   1118: 'GCU_ALARM_WORD_08_BIT_14', class GCU Alarms, trigger "60_Alarm_Data_GCU_ALARM_WORD_08" bit 6
   1119: 'GCU_ALARM_WORD_08_BIT_15', class GCU Alarms, trigger "60_Alarm_Data_GCU_ALARM_WORD_08" bit 7
   1120: 'GCU_ALARM_WORD_08_BIT_0', class GCU Alarms, trigger "60_Alarm_Data_GCU_ALARM_WORD_08" bit 8
   1121: 'GCU_ALARM_WORD_08_BIT_1', class GCU Alarms, trigger "60_Alarm_Data_GCU_ALARM_WORD_08" bit 9
   1122: 'GCU_ALARM_WORD_08_BIT_2', class GCU Alarms, trigger "60_Alarm_Data_GCU_ALARM_WORD_08" bit 10
   1123: 'GCU_ALARM_WORD_08_BIT_3', class GCU Alarms, trigger "60_Alarm_Data_GCU_ALARM_WORD_08" bit 11
   1124: 'GCU_ALARM_WORD_08_BIT_4', class GCU Alarms, trigger "60_Alarm_Data_GCU_ALARM_WORD_08" bit 12
   1125: 'GCU_ALARM_WORD_08_BIT_5', class GCU Alarms, trigger "60_Alarm_Data_GCU_ALARM_WORD_08" bit 13
   1126: 'GCU_ALARM_WORD_08_BIT_6', class GCU Alarms, trigger "60_Alarm_Data_GCU_ALARM_WORD_08" bit 14
   1127: 'GCU_ALARM_WORD_08_BIT_7', class GCU Alarms, trigger "60_Alarm_Data_GCU_ALARM_WORD_08" bit 15
   1128: 'GCU_ALARM_WORD_09_BIT_8', class GCU Alarms, trigger "60_Alarm_Data_GCU_ALARM_WORD_09" bit 0
   1129: 'GCU_ALARM_WORD_09_BIT_9', class GCU Alarms, trigger "60_Alarm_Data_GCU_ALARM_WORD_09" bit 1
   1130: 'GCU_ALARM_WORD_09_BIT_10', class GCU Alarms, trigger "60_Alarm_Data_GCU_ALARM_WORD_09" bit 2
   1131: 'GCU_ALARM_WORD_09_BIT_11', class GCU Alarms, trigger "60_Alarm_Data_GCU_ALARM_WORD_09" bit 3
   1132: 'GCU_ALARM_WORD_09_BIT_12', class GCU Alarms, trigger "60_Alarm_Data_GCU_ALARM_WORD_09" bit 4
   1133: 'GCU_ALARM_WORD_09_BIT_13', class GCU Alarms, trigger "60_Alarm_Data_GCU_ALARM_WORD_09" bit 5
   1134: 'GCU_ALARM_WORD_09_BIT_14', class GCU Alarms, trigger "60_Alarm_Data_GCU_ALARM_WORD_09" bit 6
   1135: 'GCU_ALARM_WORD_09_BIT_15', class GCU Alarms, trigger "60_Alarm_Data_GCU_ALARM_WORD_09" bit 7
   1136: 'GCU_ALARM_WORD_09_BIT_0', class GCU Alarms, trigger "60_Alarm_Data_GCU_ALARM_WORD_09" bit 8
   1137: 'GCU_ALARM_WORD_09_BIT_1', class GCU Alarms, trigger "60_Alarm_Data_GCU_ALARM_WORD_09" bit 9
   1138: 'GCU_ALARM_WORD_09_BIT_2', class GCU Alarms, trigger "60_Alarm_Data_GCU_ALARM_WORD_09" bit 10
   1139: 'GCU_ALARM_WORD_09_BIT_3', class GCU Alarms, trigger "60_Alarm_Data_GCU_ALARM_WORD_09" bit 11
   1140: 'GCU_ALARM_WORD_09_BIT_4', class GCU Alarms, trigger "60_Alarm_Data_GCU_ALARM_WORD_09" bit 12
   1141: 'GCU_ALARM_WORD_09_BIT_5', class GCU Alarms, trigger "60_Alarm_Data_GCU_ALARM_WORD_09" bit 13
   1142: 'GCU_ALARM_WORD_09_BIT_6', class GCU Alarms, trigger "60_Alarm_Data_GCU_ALARM_WORD_09" bit 14
   1143: 'GCU_ALARM_WORD_09_BIT_7', class GCU Alarms, trigger "60_Alarm_Data_GCU_ALARM_WORD_09" bit 15
   1144: 'PIT-358 FRESH WATER INLET PRESSURE', class GCU Warnings, trigger "62_Warning_Data_GCU_WARNING_WORD_01" bit 0
   1145: 'GCU_WARNING_WORD_01_BIT_9', class GCU Warnings, trigger "62_Warning_Data_GCU_WARNING_WORD_01" bit 1
   1146: 'GCU_WARNING_WORD_01_BIT_10', class GCU Warnings, trigger "62_Warning_Data_GCU_WARNING_WORD_01" bit 2
   1147: 'GCU_WARNING_WORD_01_BIT_11', class GCU Warnings, trigger "62_Warning_Data_GCU_WARNING_WORD_01" bit 3
   1148: 'GCU_WARNING_WORD_01_BIT_12', class GCU Warnings, trigger "62_Warning_Data_GCU_WARNING_WORD_01" bit 4
   1149: 'GCU_WARNING_WORD_01_BIT_13', class GCU Warnings, trigger "62_Warning_Data_GCU_WARNING_WORD_01" bit 5
   1150: 'GCU_WARNING_WORD_01_BIT_14', class GCU Warnings, trigger "62_Warning_Data_GCU_WARNING_WORD_01" bit 6
   1151: 'GCU_WARNING_WORD_01_BIT_15', class GCU Warnings, trigger "62_Warning_Data_GCU_WARNING_WORD_01" bit 7
   1152: 'PIT-348 CSW PRESSURE - OUT OF RANGE', class GCU Warnings, trigger "62_Warning_Data_GCU_WARNING_WORD_01" bit 8
   1153: 'LIT-304 LIQUID LEVEL - OUT OF RANGE', class GCU Warnings, trigger "62_Warning_Data_GCU_WARNING_WORD_01" bit 9
   1154: 'TIT-406 GAS TO DECK (OUTLET) TEMP - OUT OF RANGE', class GCU Warnings, trigger "62_Warning_Data_GCU_WARNING_WORD_01" bit 10
   1155: 'TIT-408 FRESH WATER COOLING TEMP - OUT OF RANGE', class GCU Warnings, trigger "62_Warning_Data_GCU_WARNING_WORD_01" bit 11
   1156: 'TIT-002 PGC DISCHARGE (OUTLET) TEMP - OUT OF RANGE', class GCU Warnings, trigger "62_Warning_Data_GCU_WARNING_WORD_01" bit 12
   1157: 'PIT-002 PGC DISCHARGE (OUTLET) PRESSURE - OUT OF RANGE', class GCU Warnings, trigger "62_Warning_Data_GCU_WARNING_WORD_01" bit 13
   1158: 'PIT-353 RECIRCULATION FRESH WATER PRESSURE - OUT OF RANGE', class GCU Warnings, trigger "62_Warning_Data_GCU_WARNING_WORD_01" bit 14
   1159: 'PIT-416 GAS TO DECK PRESSURE - OUT OF RANGE', class GCU Warnings, trigger "62_Warning_Data_GCU_WARNING_WORD_01" bit 15
   1160: 'PIT-002 - HIGH', class GCU Warnings, trigger "62_Warning_Data_GCU_WARNING_WORD_02" bit 0
   1161: 'PIT-353 FRESH WATER COOLING TO GCU - LOW', class GCU Warnings, trigger "62_Warning_Data_GCU_WARNING_WORD_02" bit 1
   1162: 'PIT-353 FRESH WATER COOLING TO GCU - HIGH', class GCU Warnings, trigger "62_Warning_Data_GCU_WARNING_WORD_02" bit 2
   1163: 'PIT-416 PROCESS GAS TO DECK PRESSURE - LOW', class GCU Warnings, trigger "62_Warning_Data_GCU_WARNING_WORD_02" bit 3
   1164: 'PIT-416 PROCESS GAS TO DECK PRESSURE - HIGH', class GCU Warnings, trigger "62_Warning_Data_GCU_WARNING_WORD_02" bit 4
   1165: 'PIT-358 BOOSTER FRESH WATER FILL PRESSURE - LOW', class GCU Warnings, trigger "62_Warning_Data_GCU_WARNING_WORD_02" bit 5
   1166: 'PIT-358 BOOSTER FRESH WATER FILL PRESSURE - HIGH', class GCU Warnings, trigger "62_Warning_Data_GCU_WARNING_WORD_02" bit 6
   1167: 'FS-350 FRESH WATER COOLING FLOW SWITCH - LOW FLOW5', class GCU Warnings, trigger "62_Warning_Data_GCU_WARNING_WORD_02" bit 7
   1168: 'CHECK PIT-348 COOLING SEAWATER PRESSURE', class GCU Warnings, trigger "62_Warning_Data_GCU_WARNING_WORD_02" bit 8
   1169: 'CHECK PIT-348 LOW COOLING SEAWATER PRESSURE', class GCU Warnings, trigger "62_Warning_Data_GCU_WARNING_WORD_02" bit 9
   1170: 'CHECK PIT-348 HIGH COOLING SEAWATER PRESSURE', class GCU Warnings, trigger "62_Warning_Data_GCU_WARNING_WORD_02" bit 10
   1171: 'CHECK LIT-304 GCU TANK LEVEL - HIGH', class GCU Warnings, trigger "62_Warning_Data_GCU_WARNING_WORD_02" bit 11
   1172: 'LIT-304 GCU LIQUID LEVEL - LOW', class GCU Warnings, trigger "62_Warning_Data_GCU_WARNING_WORD_02" bit 12
   1173: 'TIT-406 PROCESS GAS TO DECK TEMPERATURE - HIGH TEMP', class GCU Warnings, trigger "62_Warning_Data_GCU_WARNING_WORD_02" bit 13
   1174: 'TIT-408 FRESH WATER COOLING TO GCU TEMPERATURE - HIGH TEMP', class GCU Warnings, trigger "62_Warning_Data_GCU_WARNING_WORD_02" bit 14
   1175: 'CHECK TIT-002 PGC DISCHARGE (OUTLET) TEMPERATURE', class GCU Warnings, trigger "62_Warning_Data_GCU_WARNING_WORD_02" bit 15
   1176: 'GCU_WARNING', class GCU Warnings, trigger "62_Warning_Data_GCU_WARNING_WORD_03" bit 0
   1177: 'GCU_WARNING', class GCU Warnings, trigger "62_Warning_Data_GCU_WARNING_WORD_03" bit 1
   1178: 'GCU_WARNING', class GCU Warnings, trigger "62_Warning_Data_GCU_WARNING_WORD_03" bit 2
   1179: 'GCU_WARNING', class GCU Warnings, trigger "62_Warning_Data_GCU_WARNING_WORD_03" bit 3
   1180: 'GCU_WARNING', class GCU Warnings, trigger "62_Warning_Data_GCU_WARNING_WORD_03" bit 4
   1181: 'GCU_WARNING', class GCU Warnings, trigger "62_Warning_Data_GCU_WARNING_WORD_03" bit 5
   1182: 'GCU_WARNING', class GCU Warnings, trigger "62_Warning_Data_GCU_WARNING_WORD_03" bit 6
   1183: 'GCU_WARNING', class GCU Warnings, trigger "62_Warning_Data_GCU_WARNING_WORD_03" bit 7
   1184: 'LS-303 GCU LIQUID LEVEL - LOW', class GCU Warnings, trigger "62_Warning_Data_GCU_WARNING_WORD_03" bit 8
   1185: 'GCU_WARNING_WORD_03_BIT_1', class GCU Warnings, trigger "62_Warning_Data_GCU_WARNING_WORD_03" bit 9
   1186: 'GCU E-400 - FAULT', class GCU Warnings, trigger "62_Warning_Data_GCU_WARNING_WORD_03" bit 10
   1187: 'TIT-408 FRESH WATER COOLING TO GCU TEMPERATURE - HIGH HIGH TEMP', class GCU Warnings, trigger "62_Warning_Data_GCU_WARNING_WORD_03" bit 11
   1188: 'TIT-406 PROCESS GAS TO DECK TEMPERATURE - HIGH HIGH TEMP', class GCU Warnings, trigger "62_Warning_Data_GCU_WARNING_WORD_03" bit 12
   1189: 'GCU_WARNING_WORD_03_BIT_5', class GCU Warnings, trigger "62_Warning_Data_GCU_WARNING_WORD_03" bit 13
   1190: 'GCU_WARNING_WORD_03_BIT_6', class GCU Warnings, trigger "62_Warning_Data_GCU_WARNING_WORD_03" bit 14
   1191: 'GCU_WARNING_WORD_03_BIT_7', class GCU Warnings, trigger "62_Warning_Data_GCU_WARNING_WORD_03" bit 15
   1192: 'GCU_WARNING_WORD_04_BIT_8', class GCU Warnings, trigger "62_Warning_Data_GCU_WARNING_WORD_04" bit 0
   1193: 'GCU_WARNING_WORD_04_BIT_9', class GCU Warnings, trigger "62_Warning_Data_GCU_WARNING_WORD_04" bit 1
   1194: 'GCU_WARNING_WORD_04_BIT_10', class GCU Warnings, trigger "62_Warning_Data_GCU_WARNING_WORD_04" bit 2
   1195: 'GCU_WARNING_WORD_04_BIT_11', class GCU Warnings, trigger "62_Warning_Data_GCU_WARNING_WORD_04" bit 3
   1196: 'GCU_WARNING_WORD_04_BIT_12', class GCU Warnings, trigger "62_Warning_Data_GCU_WARNING_WORD_04" bit 4
   1197: 'GCU_WARNING_WORD_04_BIT_13', class GCU Warnings, trigger "62_Warning_Data_GCU_WARNING_WORD_04" bit 5
   1198: 'GCU_WARNING_WORD_04_BIT_14', class GCU Warnings, trigger "62_Warning_Data_GCU_WARNING_WORD_04" bit 6
   1199: 'GCU_WARNING_WORD_04_BIT_15', class GCU Warnings, trigger "62_Warning_Data_GCU_WARNING_WORD_04" bit 7
   1200: 'GCU_WARNING_WORD_04_BIT_0', class GCU Warnings, trigger "62_Warning_Data_GCU_WARNING_WORD_04" bit 8
   1201: 'GCU_WARNING_WORD_04_BIT_1', class GCU Warnings, trigger "62_Warning_Data_GCU_WARNING_WORD_04" bit 9
   1202: 'GCU_WARNING_WORD_04_BIT_2', class GCU Warnings, trigger "62_Warning_Data_GCU_WARNING_WORD_04" bit 10
   1203: 'GCU_WARNING_WORD_04_BIT_3', class GCU Warnings, trigger "62_Warning_Data_GCU_WARNING_WORD_04" bit 11
   1204: 'GCU_WARNING_WORD_04_BIT_4', class GCU Warnings, trigger "62_Warning_Data_GCU_WARNING_WORD_04" bit 12
   1205: 'GCU_WARNING_WORD_04_BIT_5', class GCU Warnings, trigger "62_Warning_Data_GCU_WARNING_WORD_04" bit 13
   1206: 'GCU_WARNING_WORD_04_BIT_6', class GCU Warnings, trigger "62_Warning_Data_GCU_WARNING_WORD_04" bit 14
   1207: 'GCU_WARNING_WORD_04_BIT_7', class GCU Warnings, trigger "62_Warning_Data_GCU_WARNING_WORD_04" bit 15
   1208: 'GCU_WARNING_WORD_05_BIT_8', class GCU Warnings, trigger "62_Warning_Data_GCU_WARNING_WORD_05" bit 0
   1209: 'GCU_WARNING_WORD_05_BIT_9', class GCU Warnings, trigger "62_Warning_Data_GCU_WARNING_WORD_05" bit 1
   1210: 'GCU_WARNING_WORD_05_BIT_10', class GCU Warnings, trigger "62_Warning_Data_GCU_WARNING_WORD_05" bit 2
   1211: 'GCU_WARNING_WORD_05_BIT_11', class GCU Warnings, trigger "62_Warning_Data_GCU_WARNING_WORD_05" bit 3
   1212: 'GCU_WARNING_WORD_05_BIT_12', class GCU Warnings, trigger "62_Warning_Data_GCU_WARNING_WORD_05" bit 4
   1213: 'GCU_WARNING_WORD_05_BIT_13', class GCU Warnings, trigger "62_Warning_Data_GCU_WARNING_WORD_05" bit 5
   1214: 'GCU_WARNING_WORD_05_BIT_14', class GCU Warnings, trigger "62_Warning_Data_GCU_WARNING_WORD_05" bit 6
   1215: 'GCU_WARNING_WORD_05_BIT_15', class GCU Warnings, trigger "62_Warning_Data_GCU_WARNING_WORD_05" bit 7
   1216: 'GCU_WARNING_WORD_05_BIT_0', class GCU Warnings, trigger "62_Warning_Data_GCU_WARNING_WORD_05" bit 8
   1217: 'GCU_WARNING_WORD_05_BIT_1', class GCU Warnings, trigger "62_Warning_Data_GCU_WARNING_WORD_05" bit 9
   1218: 'GCU_WARNING_WORD_05_BIT_2', class GCU Warnings, trigger "62_Warning_Data_GCU_WARNING_WORD_05" bit 10
   1219: 'GCU_WARNING_WORD_05_BIT_3', class GCU Warnings, trigger "62_Warning_Data_GCU_WARNING_WORD_05" bit 11
   1220: 'GCU_WARNING_WORD_05_BIT_4', class GCU Warnings, trigger "62_Warning_Data_GCU_WARNING_WORD_05" bit 12
   1221: 'GCU_WARNING_WORD_05_BIT_5', class GCU Warnings, trigger "62_Warning_Data_GCU_WARNING_WORD_05" bit 13
   1222: 'GCU_WARNING_WORD_05_BIT_6', class GCU Warnings, trigger "62_Warning_Data_GCU_WARNING_WORD_05" bit 14
   1223: 'GCU_WARNING_WORD_05_BIT_7', class GCU Warnings, trigger "62_Warning_Data_GCU_WARNING_WORD_05" bit 15
   1224: 'GCU_WARNING_WORD_06_BIT_8', class GCU Warnings, trigger "62_Warning_Data_GCU_WARNING_WORD_06" bit 0
   1225: 'GCU_WARNING_WORD_06_BIT_9', class GCU Warnings, trigger "62_Warning_Data_GCU_WARNING_WORD_06" bit 1
   1226: 'GCU_WARNING_WORD_06_BIT_10', class GCU Warnings, trigger "62_Warning_Data_GCU_WARNING_WORD_06" bit 2
   1227: 'GCU_WARNING_WORD_06_BIT_11', class GCU Warnings, trigger "62_Warning_Data_GCU_WARNING_WORD_06" bit 3
   1228: 'GCU_WARNING_WORD_06_BIT_12', class GCU Warnings, trigger "62_Warning_Data_GCU_WARNING_WORD_06" bit 4
   1229: 'GCU_WARNING_WORD_06_BIT_13', class GCU Warnings, trigger "62_Warning_Data_GCU_WARNING_WORD_06" bit 5
   1230: 'GCU_WARNING_WORD_06_BIT_14', class GCU Warnings, trigger "62_Warning_Data_GCU_WARNING_WORD_06" bit 6
   1231: 'GCU_WARNING_WORD_06_BIT_15', class GCU Warnings, trigger "62_Warning_Data_GCU_WARNING_WORD_06" bit 7
   1232: 'GCU_WARNING_WORD_06_BIT_0', class GCU Warnings, trigger "62_Warning_Data_GCU_WARNING_WORD_06" bit 8
   1233: 'GCU_WARNING_WORD_06_BIT_1', class GCU Warnings, trigger "62_Warning_Data_GCU_WARNING_WORD_06" bit 9
   1234: 'GCU_WARNING_WORD_06_BIT_2', class GCU Warnings, trigger "62_Warning_Data_GCU_WARNING_WORD_06" bit 10
   1235: 'GCU_WARNING_WORD_06_BIT_3', class GCU Warnings, trigger "62_Warning_Data_GCU_WARNING_WORD_06" bit 11
   1236: 'GCU_WARNING_WORD_06_BIT_4', class GCU Warnings, trigger "62_Warning_Data_GCU_WARNING_WORD_06" bit 12
   1237: 'GCU_WARNING_WORD_06_BIT_5', class GCU Warnings, trigger "62_Warning_Data_GCU_WARNING_WORD_06" bit 13
   1238: 'GCU_WARNING_WORD_06_BIT_6', class GCU Warnings, trigger "62_Warning_Data_GCU_WARNING_WORD_06" bit 14
   1239: 'GCU_WARNING_WORD_06_BIT_7', class GCU Warnings, trigger "62_Warning_Data_GCU_WARNING_WORD_06" bit 15
   1240: 'GCU_WARNING_WORD_07_BIT_8', class GCU Warnings, trigger "62_Warning_Data_GCU_WARNING_WORD_07" bit 0
   1241: 'GCU_WARNING_WORD_07_BIT_9', class GCU Warnings, trigger "62_Warning_Data_GCU_WARNING_WORD_07" bit 1
   1242: 'GCU_WARNING_WORD_07_BIT_10', class GCU Warnings, trigger "62_Warning_Data_GCU_WARNING_WORD_07" bit 2
   1243: 'GCU_WARNING_WORD_07_BIT_11', class GCU Warnings, trigger "62_Warning_Data_GCU_WARNING_WORD_07" bit 3
   1244: 'GCU_WARNING_WORD_07_BIT_12', class GCU Warnings, trigger "62_Warning_Data_GCU_WARNING_WORD_07" bit 4
   1245: 'GCU_WARNING_WORD_07_BIT_13', class GCU Warnings, trigger "62_Warning_Data_GCU_WARNING_WORD_07" bit 5
   1246: 'GCU_WARNING_WORD_07_BIT_14', class GCU Warnings, trigger "62_Warning_Data_GCU_WARNING_WORD_07" bit 6
   1247: 'GCU_WARNING_WORD_07_BIT_15', class GCU Warnings, trigger "62_Warning_Data_GCU_WARNING_WORD_07" bit 7
   1248: 'GCU_WARNING_WORD_07_BIT_0', class GCU Warnings, trigger "62_Warning_Data_GCU_WARNING_WORD_07" bit 8
   1249: 'GCU_WARNING_WORD_07_BIT_1', class GCU Warnings, trigger "62_Warning_Data_GCU_WARNING_WORD_07" bit 9
   1250: 'GCU_WARNING_WORD_07_BIT_2', class GCU Warnings, trigger "62_Warning_Data_GCU_WARNING_WORD_07" bit 10
   1251: 'GCU_WARNING_WORD_07_BIT_3', class GCU Warnings, trigger "62_Warning_Data_GCU_WARNING_WORD_07" bit 11
   1252: 'GCU_WARNING_WORD_07_BIT_4', class GCU Warnings, trigger "62_Warning_Data_GCU_WARNING_WORD_07" bit 12
   1253: 'GCU_WARNING_WORD_07_BIT_5', class GCU Warnings, trigger "62_Warning_Data_GCU_WARNING_WORD_07" bit 13
   1254: 'GCU_WARNING_WORD_07_BIT_6', class GCU Warnings, trigger "62_Warning_Data_GCU_WARNING_WORD_07" bit 14
   1255: 'GCU_WARNING_WORD_07_BIT_7', class GCU Warnings, trigger "62_Warning_Data_GCU_WARNING_WORD_07" bit 15
   1256: 'GCU_WARNING_WORD_08_BIT_8', class GCU Warnings, trigger "62_Warning_Data_GCU_WARNING_WORD_08" bit 0
   1257: 'GCU_WARNING_WORD_08_BIT_9', class GCU Warnings, trigger "62_Warning_Data_GCU_WARNING_WORD_08" bit 1
   1258: 'GCU_WARNING_WORD_08_BIT_10', class GCU Warnings, trigger "62_Warning_Data_GCU_WARNING_WORD_08" bit 2
   1259: 'GCU_WARNING_WORD_08_BIT_11', class GCU Warnings, trigger "62_Warning_Data_GCU_WARNING_WORD_08" bit 3
   1260: 'GCU_WARNING_WORD_08_BIT_12', class GCU Warnings, trigger "62_Warning_Data_GCU_WARNING_WORD_08" bit 4
   1261: 'GCU_WARNING_WORD_08_BIT_13', class GCU Warnings, trigger "62_Warning_Data_GCU_WARNING_WORD_08" bit 5
   1262: 'GCU_WARNING_WORD_08_BIT_14', class GCU Warnings, trigger "62_Warning_Data_GCU_WARNING_WORD_08" bit 6
   1263: 'GCU_WARNING_WORD_08_BIT_15', class GCU Warnings, trigger "62_Warning_Data_GCU_WARNING_WORD_08" bit 7
   1264: 'GCU_WARNING_WORD_08_BIT_0', class GCU Warnings, trigger "62_Warning_Data_GCU_WARNING_WORD_08" bit 8
   1265: 'GCU_WARNING_WORD_08_BIT_1', class GCU Warnings, trigger "62_Warning_Data_GCU_WARNING_WORD_08" bit 9
   1266: 'GCU_WARNING_WORD_08_BIT_2', class GCU Warnings, trigger "62_Warning_Data_GCU_WARNING_WORD_08" bit 10
   1267: 'GCU_WARNING_WORD_08_BIT_3', class GCU Warnings, trigger "62_Warning_Data_GCU_WARNING_WORD_08" bit 11
   1268: 'GCU_WARNING_WORD_08_BIT_4', class GCU Warnings, trigger "62_Warning_Data_GCU_WARNING_WORD_08" bit 12
   1269: 'GCU_WARNING_WORD_08_BIT_5', class GCU Warnings, trigger "62_Warning_Data_GCU_WARNING_WORD_08" bit 13
   1270: 'GCU_WARNING_WORD_08_BIT_6', class GCU Warnings, trigger "62_Warning_Data_GCU_WARNING_WORD_08" bit 14
   1271: 'GCU_WARNING_WORD_08_BIT_7', class GCU Warnings, trigger "62_Warning_Data_GCU_WARNING_WORD_08" bit 15
   1272: 'GCU_WARNING_WORD_09_BIT_8', class GCU Warnings, trigger "62_Warning_Data_GCU_WARNING_WORD_09" bit 0
   1273: 'GCU_WARNING_WORD_09_BIT_9', class GCU Warnings, trigger "62_Warning_Data_GCU_WARNING_WORD_09" bit 1
   1274: 'GCU_WARNING_WORD_09_BIT_10', class GCU Warnings, trigger "62_Warning_Data_GCU_WARNING_WORD_09" bit 2
   1275: 'GCU_WARNING_WORD_09_BIT_11', class GCU Warnings, trigger "62_Warning_Data_GCU_WARNING_WORD_09" bit 3
   1276: 'GCU_WARNING_WORD_09_BIT_12', class GCU Warnings, trigger "62_Warning_Data_GCU_WARNING_WORD_09" bit 4
   1277: 'GCU_WARNING_WORD_09_BIT_13', class GCU Warnings, trigger "62_Warning_Data_GCU_WARNING_WORD_09" bit 5
   1278: 'GCU_WARNING_WORD_09_BIT_14', class GCU Warnings, trigger "62_Warning_Data_GCU_WARNING_WORD_09" bit 6
   1279: 'GCU_WARNING_WORD_09_BIT_15', class GCU Warnings, trigger "62_Warning_Data_GCU_WARNING_WORD_09" bit 7
   1280: 'GCU_WARNING_WORD_09_BIT_0', class GCU Warnings, trigger "62_Warning_Data_GCU_WARNING_WORD_09" bit 8
   1281: 'GCU_WARNING_WORD_09_BIT_1', class GCU Warnings, trigger "62_Warning_Data_GCU_WARNING_WORD_09" bit 9
   1282: 'GCU_WARNING_WORD_09_BIT_2', class GCU Warnings, trigger "62_Warning_Data_GCU_WARNING_WORD_09" bit 10
   1283: 'GCU_WARNING_WORD_09_BIT_3', class GCU Warnings, trigger "62_Warning_Data_GCU_WARNING_WORD_09" bit 11
   1284: 'GCU_WARNING_WORD_09_BIT_4', class GCU Warnings, trigger "62_Warning_Data_GCU_WARNING_WORD_09" bit 12
   1285: 'GCU_WARNING_WORD_09_BIT_5', class GCU Warnings, trigger "62_Warning_Data_GCU_WARNING_WORD_09" bit 13
   1286: 'GCU_WARNING_WORD_09_BIT_6', class GCU Warnings, trigger "62_Warning_Data_GCU_WARNING_WORD_09" bit 14
   1287: 'GCU_WARNING_WORD_09_BIT_7', class GCU Warnings, trigger "62_Warning_Data_GCU_WARNING_WORD_09" bit 15
   2000: 'FIT-418 2 PORT USD FLOW - LOW LOW', class Tank Control Alarms, trigger "2060_Alarm_Data_BTCS_ALARM_WORD_01" bit 0
   2001: 'FIT-418 2 PORT USD FLOW - HIGH HIGH', class Tank Control Alarms, trigger "2060_Alarm_Data_BTCS_ALARM_WORD_01" bit 1
   2002: 'FIT-420 2 PORT MBG FLOW - LOW LOW', class Tank Control Alarms, trigger "2060_Alarm_Data_BTCS_ALARM_WORD_01" bit 2
   2003: 'FIT-420 2 PORT MBG FLOW - HIGH HIGH', class Tank Control Alarms, trigger "2060_Alarm_Data_BTCS_ALARM_WORD_01" bit 3
   2004: 'FIT-417 2 STARBOARD USD FLOW - LOW LOW', class Tank Control Alarms, trigger "2060_Alarm_Data_BTCS_ALARM_WORD_01" bit 4
   2005: 'FIT-417 2 STARBOARD USD FLOW - HIGH HIGH', class Tank Control Alarms, trigger "2060_Alarm_Data_BTCS_ALARM_WORD_01" bit 5
   2006: 'FIT-419 2 STARBOARD MBG FLOW - LOW LOW', class Tank Control Alarms, trigger "2060_Alarm_Data_BTCS_ALARM_WORD_01" bit 6
   2007: 'FIT-419 2 STARBOARD MBG FLOW - HIGH HIGH', class Tank Control Alarms, trigger "2060_Alarm_Data_BTCS_ALARM_WORD_01" bit 7
   2008: 'CV-442 2 PORT GAS to TANK VALVE FAULT', class Tank Control Alarms, trigger "2060_Alarm_Data_BTCS_ALARM_WORD_01" bit 8
   2009: 'CV-441 2 STARBOARD GAS to TANK VALVE FAULT', class Tank Control Alarms, trigger "2060_Alarm_Data_BTCS_ALARM_WORD_01" bit 9
   2010: 'TIT-436 2 PORT BWT TEMP - HIGH HIGH', class Tank Control Alarms, trigger "2060_Alarm_Data_BTCS_ALARM_WORD_01" bit 10
   2011: 'TIT-436 2 STARBOARD BWT TEMP - HIGH HIGH', class Tank Control Alarms, trigger "2060_Alarm_Data_BTCS_ALARM_WORD_01" bit 11
   2012: 'LS-425 2 PORT LEVEL - HIGH HIGH', class Tank Control Alarms, trigger "2060_Alarm_Data_BTCS_ALARM_WORD_01" bit 12
   2013: 'LS-425 2 STARBOARD LEVEL - HIGH HIGH', class Tank Control Alarms, trigger "2060_Alarm_Data_BTCS_ALARM_WORD_01" bit 13
   2014: 'PS-436 2 BALLAST TANK PRESSURE - HIGH', class Tank Control Alarms, trigger "2060_Alarm_Data_BTCS_ALARM_WORD_01" bit 14
   2015: '600-TX-433 APT O2 MONITOR - LOW', class Tank Control Alarms, trigger "2060_Alarm_Data_BTCS_ALARM_WORD_01" bit 15
   2016: 'CV422 FPT GAS to TANK VALVE FAULT', class Tank Control Alarms, trigger "2060_Alarm_Data_BTCS_ALARM_WORD_02" bit 0
   2017: 'CV422 1 PORT GAS to TANK VALVE FAULT', class Tank Control Alarms, trigger "2060_Alarm_Data_BTCS_ALARM_WORD_02" bit 1
   2018: 'CV421 1 STARBOARD GAS to TANK VALVE FAULT', class Tank Control Alarms, trigger "2060_Alarm_Data_BTCS_ALARM_WORD_02" bit 2
   2019: 'CV422 3 PORT GAS to TANK VALVE FAULT', class Tank Control Alarms, trigger "2060_Alarm_Data_BTCS_ALARM_WORD_02" bit 3
   2020: 'CV421 3 STARBOARD GAS to TANK VALVE FAULT', class Tank Control Alarms, trigger "2060_Alarm_Data_BTCS_ALARM_WORD_02" bit 4
   2021: 'CV422 4 PORT GAS to TANK VALVE FAULT', class Tank Control Alarms, trigger "2060_Alarm_Data_BTCS_ALARM_WORD_02" bit 5
   2022: 'CV421 4 STARBOARD GAS to TANK VALVE FAULT', class Tank Control Alarms, trigger "2060_Alarm_Data_BTCS_ALARM_WORD_02" bit 6
   2023: 'CV422 5 PORT GAS to TANK VALVE FAULT', class Tank Control Alarms, trigger "2060_Alarm_Data_BTCS_ALARM_WORD_02" bit 7
   2024: 'PIT-415 2 PORT DECK IG PRESSURE - LOW LOW', class Tank Control Alarms, trigger "2060_Alarm_Data_BTCS_ALARM_WORD_02" bit 8
   2025: 'PIT-415 2 PORT DECK IG PRESSURE - HIGH HIGH', class Tank Control Alarms, trigger "2060_Alarm_Data_BTCS_ALARM_WORD_02" bit 9
   2026: 'PIT-415 2 STARBOARD DECK IG PRESSURE - LOW LOW', class Tank Control Alarms, trigger "2060_Alarm_Data_BTCS_ALARM_WORD_02" bit 10
   2027: 'PIT-415 2 STARBOARD DECK IG PRESSURE - HIGH HIGH', class Tank Control Alarms, trigger "2060_Alarm_Data_BTCS_ALARM_WORD_02" bit 11
   2028: 'PIT-424 2 PORT TANK PRESSURE - LOW LOW', class Tank Control Alarms, trigger "2060_Alarm_Data_BTCS_ALARM_WORD_02" bit 12
   2029: 'PIT-424 2 PORT TANK PRESSURE - HIGH HIGH', class Tank Control Alarms, trigger "2060_Alarm_Data_BTCS_ALARM_WORD_02" bit 13
   2030: 'PIT-424 2 STARBOARD TANK PRESSURE - LOW LOW', class Tank Control Alarms, trigger "2060_Alarm_Data_BTCS_ALARM_WORD_02" bit 14
   2031: 'PIT-424 2 STARBOARD TANK PRESSURE - HIGH HIGH', class Tank Control Alarms, trigger "2060_Alarm_Data_BTCS_ALARM_WORD_02" bit 15
   2128: 'FIT-418 2 PORT USD FLOW - LOW', class Tank Control Warnings, trigger "2062_Warning_Data_BTCS_WARNING_WORD_01" bit 0
   2129: 'FIT-418 2 PORT USD FLOW - HIGH', class Tank Control Warnings, trigger "2062_Warning_Data_BTCS_WARNING_WORD_01" bit 1
   2130: 'FIT-420 2 PORT MBG FLOW - LOW', class Tank Control Warnings, trigger "2062_Warning_Data_BTCS_WARNING_WORD_01" bit 2
   2131: 'FIT-420 2 PORT MBG FLOW - HIGH', class Tank Control Warnings, trigger "2062_Warning_Data_BTCS_WARNING_WORD_01" bit 3
   2132: 'FIT-417 2 STARBOARD USD FLOW - LOW', class Tank Control Warnings, trigger "2062_Warning_Data_BTCS_WARNING_WORD_01" bit 4
   2133: 'FIT-417 2 STARBOARD USD FLOW - HIGH', class Tank Control Warnings, trigger "2062_Warning_Data_BTCS_WARNING_WORD_01" bit 5
   2134: 'FIT-419 2 STARBOARD MBG FLOW - LOW', class Tank Control Warnings, trigger "2062_Warning_Data_BTCS_WARNING_WORD_01" bit 6
   2135: 'FIT-419 2 STARBOARD MBG FLOW - HIGH', class Tank Control Warnings, trigger "2062_Warning_Data_BTCS_WARNING_WORD_01" bit 7
   2136: '600-TX-433 APT O2 MONITOR - LOW', class Tank Control Warnings, trigger "2062_Warning_Data_BTCS_WARNING_WORD_01" bit 8
   2137: '600-TX-433 APT O2 MONITOR - LOW LOW', class Tank Control Warnings, trigger "2062_Warning_Data_BTCS_WARNING_WORD_01" bit 9
   2138: 'TIT-436 2 PORT BWT TEMP - HIGH', class Tank Control Warnings, trigger "2062_Warning_Data_BTCS_WARNING_WORD_01" bit 10
   2139: 'TIT-436 2 STARBOARD BWT TEMP - HIGH', class Tank Control Warnings, trigger "2062_Warning_Data_BTCS_WARNING_WORD_01" bit 11
   2140: 'BTCS_WARNING_WORD_01_BIT_4', class Tank Control Warnings, trigger "2062_Warning_Data_BTCS_WARNING_WORD_01" bit 12
   2141: 'BTCS_WARNING_WORD_01_BIT_5', class Tank Control Warnings, trigger "2062_Warning_Data_BTCS_WARNING_WORD_01" bit 13
   2142: 'BTCS_WARNING_WORD_01_BIT_6', class Tank Control Warnings, trigger "2062_Warning_Data_BTCS_WARNING_WORD_01" bit 14
   2143: 'BTCS_WARNING_WORD_01_BIT_7', class Tank Control Warnings, trigger "2062_Warning_Data_BTCS_WARNING_WORD_01" bit 15
   2144: 'TT-426 1 FOR PEACK TANK TEMPERATURE - HIGH', class Tank Control Warnings, trigger "2062_Warning_Data_BTCS_WARNING_WORD_02" bit 0
   2145: 'TT-426 1 PORT TANK TEMPERATURE - HIGH', class Tank Control Warnings, trigger "2062_Warning_Data_BTCS_WARNING_WORD_02" bit 1
   2146: 'TT-426 1 STARBOARD TANK TEMPERATURE - HIGH', class Tank Control Warnings, trigger "2062_Warning_Data_BTCS_WARNING_WORD_02" bit 2
   2147: 'TT-426 3 PORT TANK TEMPERATURE - HIGH', class Tank Control Warnings, trigger "2062_Warning_Data_BTCS_WARNING_WORD_02" bit 3
   2148: 'TT-426 3 STARBOARD TANK TEMPERATURE - HIGH', class Tank Control Warnings, trigger "2062_Warning_Data_BTCS_WARNING_WORD_02" bit 4
   2149: 'TT-426 4 PORT TANK TEMPERATURE - HIGH', class Tank Control Warnings, trigger "2062_Warning_Data_BTCS_WARNING_WORD_02" bit 5
   2150: 'TT-426 4 STARBOARD TANK TEMPERATURE - HIGH', class Tank Control Warnings, trigger "2062_Warning_Data_BTCS_WARNING_WORD_02" bit 6
   2151: 'TT-426 5 PORT TANK TEMPERATURE - HIGH', class Tank Control Warnings, trigger "2062_Warning_Data_BTCS_WARNING_WORD_02" bit 7
   2152: 'PIT-415 2 PORT DECK IG PRESSURE - LOW', class Tank Control Warnings, trigger "2062_Warning_Data_BTCS_WARNING_WORD_02" bit 8
   2153: 'PIT-415 2 PORT DECK IG PRESSURE - HIGH', class Tank Control Warnings, trigger "2062_Warning_Data_BTCS_WARNING_WORD_02" bit 9
   2154: 'PIT-415 2 STARBOARD DECK IG PRESSURE - LOW', class Tank Control Warnings, trigger "2062_Warning_Data_BTCS_WARNING_WORD_02" bit 10
   2155: 'PIT-415 STARBOARD DECK IG PRESSURE - HIGH', class Tank Control Warnings, trigger "2062_Warning_Data_BTCS_WARNING_WORD_02" bit 11
   2156: 'PIT-424 2 PORT TANK PRESSURE - LOW', class Tank Control Warnings, trigger "2062_Warning_Data_BTCS_WARNING_WORD_02" bit 12
   2157: 'PIT-424 2 PORT TANK PRESSURE - HIGH', class Tank Control Warnings, trigger "2062_Warning_Data_BTCS_WARNING_WORD_02" bit 13
   2158: 'PIT-424 2 STARBOARD TANK PRESSURE - LOW', class Tank Control Warnings, trigger "2062_Warning_Data_BTCS_WARNING_WORD_02" bit 14
   2159: 'PIT-424 2 STARBOARD TANK PRESSURE - HIGH', class Tank Control Warnings, trigger "2062_Warning_Data_BTCS_WARNING_WORD_02" bit 15
   2160: 'FIT418 1 FOR PEACK TANK USD FLOW LOW', class Tank Control Warnings, trigger "2062_Warning_Data_BTCS_WARNING_WORD_03" bit 0
   2161: 'FIT418 1 FOR PEACK TANK USD FLOW HIGH', class Tank Control Warnings, trigger "2062_Warning_Data_BTCS_WARNING_WORD_03" bit 1
   2162: 'FIT418 1 PORT TANK USD FLOW LOW', class Tank Control Warnings, trigger "2062_Warning_Data_BTCS_WARNING_WORD_03" bit 2
   2163: 'FIT418 1 PORT TANK USD FLOW HIGH', class Tank Control Warnings, trigger "2062_Warning_Data_BTCS_WARNING_WORD_03" bit 3
   2164: 'FIT417 1 STARBOARD TANK USD FLOW LOW', class Tank Control Warnings, trigger "2062_Warning_Data_BTCS_WARNING_WORD_03" bit 4
   2165: 'FIT417 1 STARBOARD TANK USD FLOW HIGH', class Tank Control Warnings, trigger "2062_Warning_Data_BTCS_WARNING_WORD_03" bit 5
   2166: 'FIT418 3 PORT TANK USD FLOW LOW', class Tank Control Warnings, trigger "2062_Warning_Data_BTCS_WARNING_WORD_03" bit 6
   2167: 'FIT418 3 PORT TANK USD FLOW HIGH', class Tank Control Warnings, trigger "2062_Warning_Data_BTCS_WARNING_WORD_03" bit 7
   2168: 'TT-426 5 STARBOARD TANK TEMPERATURE - HIGH', class Tank Control Warnings, trigger "2062_Warning_Data_BTCS_WARNING_WORD_03" bit 8
   2169: 'TT-426 6 PORT TANK TEMPERATURE - HIGH', class Tank Control Warnings, trigger "2062_Warning_Data_BTCS_WARNING_WORD_03" bit 9
   2170: 'TT-426 6 STARBOARD TANK TEMPERATURE - HIGH', class Tank Control Warnings, trigger "2062_Warning_Data_BTCS_WARNING_WORD_03" bit 10
   2171: 'TT-426 7 AFT PEACK TANK TEMPERATURE - HIGH', class Tank Control Warnings, trigger "2062_Warning_Data_BTCS_WARNING_WORD_03" bit 11
   2172: 'BTCS_WARNING_WORD_03_BIT_4', class Tank Control Warnings, trigger "2062_Warning_Data_BTCS_WARNING_WORD_03" bit 12
   2173: 'BTCS_WARNING_WORD_03_BIT_5', class Tank Control Warnings, trigger "2062_Warning_Data_BTCS_WARNING_WORD_03" bit 13
   2174: 'BTCS_WARNING_WORD_03_BIT_6', class Tank Control Warnings, trigger "2062_Warning_Data_BTCS_WARNING_WORD_03" bit 14
   2175: 'BTCS_WARNING_WORD_03_BIT_7', class Tank Control Warnings, trigger "2062_Warning_Data_BTCS_WARNING_WORD_03" bit 15
   2176: 'FIT417 5 STARBOARD TANK USD FLOW LOW', class Tank Control Warnings, trigger "2062_Warning_Data_BTCS_WARNING_WORD_04" bit 0
   2177: 'FIT417 5 STARBOARD TANK USD FLOW HIGH', class Tank Control Warnings, trigger "2062_Warning_Data_BTCS_WARNING_WORD_04" bit 1
   2178: 'FIT418 6 PORT TANK USD FLOW LOW', class Tank Control Warnings, trigger "2062_Warning_Data_BTCS_WARNING_WORD_04" bit 2
   2179: 'FIT418 6 PORT TANK USD FLOW HIGH', class Tank Control Warnings, trigger "2062_Warning_Data_BTCS_WARNING_WORD_04" bit 3
   2180: 'FIT417 6 STARBOARD TANK USD FLOW LOW', class Tank Control Warnings, trigger "2062_Warning_Data_BTCS_WARNING_WORD_04" bit 4
   2181: 'FIT417 6 STARBOARD TANK USD FLOW HIGH', class Tank Control Warnings, trigger "2062_Warning_Data_BTCS_WARNING_WORD_04" bit 5
   2182: 'FIT418 7 APT TANK USD FLOW LOW', class Tank Control Warnings, trigger "2062_Warning_Data_BTCS_WARNING_WORD_04" bit 6
   2183: 'FIT418 7 APT TANK USD FLOW HIGH', class Tank Control Warnings, trigger "2062_Warning_Data_BTCS_WARNING_WORD_04" bit 7
   2184: 'FIT417 3 STARBOARD TANK USD FLOW LOW', class Tank Control Warnings, trigger "2062_Warning_Data_BTCS_WARNING_WORD_04" bit 8
   2185: 'FIT417 3 STARBOARD TANK USD FLOW HIGH', class Tank Control Warnings, trigger "2062_Warning_Data_BTCS_WARNING_WORD_04" bit 9
   2186: 'FIT418 4 PORT TANK USD FLOW LOW', class Tank Control Warnings, trigger "2062_Warning_Data_BTCS_WARNING_WORD_04" bit 10
   2187: 'FIT418 4 PORT TANK USD FLOW HIGH', class Tank Control Warnings, trigger "2062_Warning_Data_BTCS_WARNING_WORD_04" bit 11
   2188: 'FIT417 4 STARBOARD TANK USD FLOW LOW', class Tank Control Warnings, trigger "2062_Warning_Data_BTCS_WARNING_WORD_04" bit 12
   2189: 'FIT417 4 STARBOARD TANK USD FLOW HIGH', class Tank Control Warnings, trigger "2062_Warning_Data_BTCS_WARNING_WORD_04" bit 13
   2190: 'FIT418 5 PORT TANK USD FLOW LOW', class Tank Control Warnings, trigger "2062_Warning_Data_BTCS_WARNING_WORD_04" bit 14
   2191: 'FIT418 5 PORT TANK USD FLOW HIGH', class Tank Control Warnings, trigger "2062_Warning_Data_BTCS_WARNING_WORD_04" bit 15
   2192: 'FIT419 3 STARBOARD MBG FLOW LOW', class Tank Control Warnings, trigger "2062_Warning_Data_BTCS_WARNING_WORD_05" bit 0
   2193: 'FIT419 3 STARBOARD MBG FLOW HIGH', class Tank Control Warnings, trigger "2062_Warning_Data_BTCS_WARNING_WORD_05" bit 1
   2194: 'FIT420 4 PORT MBG FLOW LOW', class Tank Control Warnings, trigger "2062_Warning_Data_BTCS_WARNING_WORD_05" bit 2
   2195: 'FIT420 4 PORT MBG FLOW HIGH', class Tank Control Warnings, trigger "2062_Warning_Data_BTCS_WARNING_WORD_05" bit 3
   2196: 'FIT419 4 STARBOARD MBG FLOW LOW', class Tank Control Warnings, trigger "2062_Warning_Data_BTCS_WARNING_WORD_05" bit 4
   2197: 'FIT419 4 STARBOARD MBG FLOW HIGH', class Tank Control Warnings, trigger "2062_Warning_Data_BTCS_WARNING_WORD_05" bit 5
   2198: 'FIT420 5 PORT MBG FLOW LOW', class Tank Control Warnings, trigger "2062_Warning_Data_BTCS_WARNING_WORD_05" bit 6
   2199: 'FIT420 5 PORT MBG FLOW HIGH', class Tank Control Warnings, trigger "2062_Warning_Data_BTCS_WARNING_WORD_05" bit 7
   2200: 'FIT420 1 FPT MBG FLOW LOW', class Tank Control Warnings, trigger "2062_Warning_Data_BTCS_WARNING_WORD_05" bit 8
   2201: 'FIT420 1 FPT MBG FLOW HIGH', class Tank Control Warnings, trigger "2062_Warning_Data_BTCS_WARNING_WORD_05" bit 9
   2202: 'FIT420 1 PORT MBG FLOW LOW', class Tank Control Warnings, trigger "2062_Warning_Data_BTCS_WARNING_WORD_05" bit 10
   2203: 'FIT420 1 PORT MBG FLOW HIGH', class Tank Control Warnings, trigger "2062_Warning_Data_BTCS_WARNING_WORD_05" bit 11
   2204: 'FIT419 1 STARBOARD MBG FLOW LOW', class Tank Control Warnings, trigger "2062_Warning_Data_BTCS_WARNING_WORD_05" bit 12
   2205: 'FIT419 1 STARBOARD MBG FLOW HIGH', class Tank Control Warnings, trigger "2062_Warning_Data_BTCS_WARNING_WORD_05" bit 13
   2206: 'FIT420 3 PORT MBG FLOW LOW', class Tank Control Warnings, trigger "2062_Warning_Data_BTCS_WARNING_WORD_05" bit 14
   2207: 'FIT420 3 PORT MBG FLOW HIGH', class Tank Control Warnings, trigger "2062_Warning_Data_BTCS_WARNING_WORD_05" bit 15
   2208: 'PT415 RIO1 DECK IG PRESSURE LOW', class Tank Control Warnings, trigger "2062_Warning_Data_BTCS_WARNING_WORD_06" bit 0
   2209: 'PT415 RIO1 DECK IG PRESSURE HIGH', class Tank Control Warnings, trigger "2062_Warning_Data_BTCS_WARNING_WORD_06" bit 1
   2210: 'PT415 RIO3 DECK IG PRESSURE LOW', class Tank Control Warnings, trigger "2062_Warning_Data_BTCS_WARNING_WORD_06" bit 2
   2211: 'PT415 RIO3 DECK IG PRESSURE HIGH', class Tank Control Warnings, trigger "2062_Warning_Data_BTCS_WARNING_WORD_06" bit 3
   2212: 'PT415 RIO4 DECK IG PRESSURE LOW', class Tank Control Warnings, trigger "2062_Warning_Data_BTCS_WARNING_WORD_06" bit 4
   2213: 'PT415 RIO4 DECK IG PRESSURE HIGH', class Tank Control Warnings, trigger "2062_Warning_Data_BTCS_WARNING_WORD_06" bit 5
   2214: 'PT415 RIO5 DECK IG PRESSURE LOW', class Tank Control Warnings, trigger "2062_Warning_Data_BTCS_WARNING_WORD_06" bit 6
   2215: 'PT415 RIO5 DECK IG PRESSURE HIGH', class Tank Control Warnings, trigger "2062_Warning_Data_BTCS_WARNING_WORD_06" bit 7
   2216: 'FIT419 5 STARBOARD MBG FLOW LOW', class Tank Control Warnings, trigger "2062_Warning_Data_BTCS_WARNING_WORD_06" bit 8
   2217: 'FIT419 5 STARBOARD MBG FLOW HIGH', class Tank Control Warnings, trigger "2062_Warning_Data_BTCS_WARNING_WORD_06" bit 9
   2218: 'FIT420 6 PORT MBG FLOW LOW', class Tank Control Warnings, trigger "2062_Warning_Data_BTCS_WARNING_WORD_06" bit 10
   2219: 'FIT420 6 PORT MBG FLOW HIGH', class Tank Control Warnings, trigger "2062_Warning_Data_BTCS_WARNING_WORD_06" bit 11
   2220: 'FIT419 6 STARBOARD MBG FLOW LOW', class Tank Control Warnings, trigger "2062_Warning_Data_BTCS_WARNING_WORD_06" bit 12
   2221: 'FIT419 6 STARBOARD MBG FLOW HIGH', class Tank Control Warnings, trigger "2062_Warning_Data_BTCS_WARNING_WORD_06" bit 13
   2222: 'FIT420 7 APT MBG FLOW LOW', class Tank Control Warnings, trigger "2062_Warning_Data_BTCS_WARNING_WORD_06" bit 14
   2223: 'FIT420 7 APT MBG FLOW HIGH', class Tank Control Warnings, trigger "2062_Warning_Data_BTCS_WARNING_WORD_06" bit 15
   2224: 'PIT424 RIO5 TANK PRESSURE LOW', class Tank Control Warnings, trigger "2062_Warning_Data_BTCS_WARNING_WORD_07" bit 0
   2225: 'PIT424 RIO5 TANK PRESSURE HIGH', class Tank Control Warnings, trigger "2062_Warning_Data_BTCS_WARNING_WORD_07" bit 1
   2226: 'PIT424 RIO6 TANK PRESSURE LOW', class Tank Control Warnings, trigger "2062_Warning_Data_BTCS_WARNING_WORD_07" bit 2
   2227: 'PIT424 RIO6 TANK PRESSURE HIGH', class Tank Control Warnings, trigger "2062_Warning_Data_BTCS_WARNING_WORD_07" bit 3
   2228: 'PIT424 RIO7 TANK PRESSURE LOW', class Tank Control Warnings, trigger "2062_Warning_Data_BTCS_WARNING_WORD_07" bit 4
   2229: 'PIT424 RIO7 TANK PRESSURE HIGH', class Tank Control Warnings, trigger "2062_Warning_Data_BTCS_WARNING_WORD_07" bit 5
   2230: 'BTCS_WARNING_WORD_07_BIT_14', class Tank Control Warnings, trigger "2062_Warning_Data_BTCS_WARNING_WORD_07" bit 6
   2231: 'BTCS_WARNING_WORD_07_BIT_15', class Tank Control Warnings, trigger "2062_Warning_Data_BTCS_WARNING_WORD_07" bit 7
   2232: 'PT415 RIO6 DECK IG PRESSURE LOW', class Tank Control Warnings, trigger "2062_Warning_Data_BTCS_WARNING_WORD_07" bit 8
   2233: 'PT415 RIO6 DECK IG PRESSURE HIGH', class Tank Control Warnings, trigger "2062_Warning_Data_BTCS_WARNING_WORD_07" bit 9
   2234: 'PIT424 RIO1 TANK PRESSURE LOW', class Tank Control Warnings, trigger "2062_Warning_Data_BTCS_WARNING_WORD_07" bit 10
   2235: 'PIT424 RIO1 TANK PRESSURE HIGH', class Tank Control Warnings, trigger "2062_Warning_Data_BTCS_WARNING_WORD_07" bit 11
   2236: 'PIT424 RIO3 TANK PRESSURE LOW', class Tank Control Warnings, trigger "2062_Warning_Data_BTCS_WARNING_WORD_07" bit 12
   2237: 'PIT424 RIO3 TANK PRESSURE HIGH', class Tank Control Warnings, trigger "2062_Warning_Data_BTCS_WARNING_WORD_07" bit 13
   2238: 'PIT424 RIO4 TANK PRESSURE LOW', class Tank Control Warnings, trigger "2062_Warning_Data_BTCS_WARNING_WORD_07" bit 14
   2239: 'PIT424 RIO4 TANK PRESSURE HIGH', class Tank Control Warnings, trigger "2062_Warning_Data_BTCS_WARNING_WORD_07" bit 15
   2240: 'LS425 4 STARBOARD TANK LEVEL HIGH HIGH', class Tank Control Warnings, trigger "2062_Warning_Data_BTCS_WARNING_WORD_08" bit 0
   2241: 'LS425 5 PORT TANK LEVEL HIGH HIGH', class Tank Control Warnings, trigger "2062_Warning_Data_BTCS_WARNING_WORD_08" bit 1
   2242: 'LS425 5 STARBOARD TANK LEVEL HIGH HIGH', class Tank Control Warnings, trigger "2062_Warning_Data_BTCS_WARNING_WORD_08" bit 2
   2243: 'LS425 6 PORT TANK LEVEL HIGH HIGH', class Tank Control Warnings, trigger "2062_Warning_Data_BTCS_WARNING_WORD_08" bit 3
   2244: 'LS425 6 STARBOARD TANK LEVEL HIGH HIGH', class Tank Control Warnings, trigger "2062_Warning_Data_BTCS_WARNING_WORD_08" bit 4
   2245: 'LS425 AP TANK LEVEL HIGH HIGH', class Tank Control Warnings, trigger "2062_Warning_Data_BTCS_WARNING_WORD_08" bit 5
   2246: 'BTCS_WARNING_WORD_08_BIT_14', class Tank Control Warnings, trigger "2062_Warning_Data_BTCS_WARNING_WORD_08" bit 6
   2247: 'LS425 FP TANK LEVEL HIGH HIGH', class Tank Control Warnings, trigger "2062_Warning_Data_BTCS_WARNING_WORD_08" bit 7
   2248: 'PT415 RIO7 DECK IG PRESSURE LOW', class Tank Control Warnings, trigger "2062_Warning_Data_BTCS_WARNING_WORD_08" bit 8
   2249: 'PT415 RIO7 DECK IG PRESSURE HIGH', class Tank Control Warnings, trigger "2062_Warning_Data_BTCS_WARNING_WORD_08" bit 9
   2250: 'LS425 1 STARBOARD TANK LEVEL HIGH HIGH', class Tank Control Warnings, trigger "2062_Warning_Data_BTCS_WARNING_WORD_08" bit 10
   2251: 'LS425 2 PORT TANK LEVEL HIGH HIGH', class Tank Control Warnings, trigger "2062_Warning_Data_BTCS_WARNING_WORD_08" bit 11
   2252: 'LS425 2 STARBOARD TANK LEVEL HIGH HIGH', class Tank Control Warnings, trigger "2062_Warning_Data_BTCS_WARNING_WORD_08" bit 12
   2253: 'LS425 3 PORT TANK LEVEL HIGH HIGH', class Tank Control Warnings, trigger "2062_Warning_Data_BTCS_WARNING_WORD_08" bit 13
   2254: 'LS425 3 STARBOARD TANK LEVEL HIGH HIGH', class Tank Control Warnings, trigger "2062_Warning_Data_BTCS_WARNING_WORD_08" bit 14
   2255: 'LS425 4 PORT TANK LEVEL HIGH HIGH', class Tank Control Warnings, trigger "2062_Warning_Data_BTCS_WARNING_WORD_08" bit 15
   2256: 'LT422 FPT TANK LEVEL HIGH', class Tank Control Warnings, trigger "2062_Warning_Data_BTCS_WARNING_WORD_09" bit 0
   2257: 'LT422 FPT TANK LEVEL LOW', class Tank Control Warnings, trigger "2062_Warning_Data_BTCS_WARNING_WORD_09" bit 1
   2258: 'LT422 1 PORT TANK LEVEL HIGH', class Tank Control Warnings, trigger "2062_Warning_Data_BTCS_WARNING_WORD_09" bit 2
   2259: 'LT422 1 PORT TANK LEVEL LOW', class Tank Control Warnings, trigger "2062_Warning_Data_BTCS_WARNING_WORD_09" bit 3
   2260: 'LT422 1 STARBOARD TANK LEVEL HIGH', class Tank Control Warnings, trigger "2062_Warning_Data_BTCS_WARNING_WORD_09" bit 4
   2261: 'LT422 1 STARBOARD TANK LEVEL LOW', class Tank Control Warnings, trigger "2062_Warning_Data_BTCS_WARNING_WORD_09" bit 5
   2262: 'LT422 2 PORT TANK LEVEL HIGH', class Tank Control Warnings, trigger "2062_Warning_Data_BTCS_WARNING_WORD_09" bit 6
   2263: 'LT422 2 PORT TANK LEVEL LOW', class Tank Control Warnings, trigger "2062_Warning_Data_BTCS_WARNING_WORD_09" bit 7
   2264: 'PS436 RIO1 TANK GROUP PRESURE HIGH HIGH', class Tank Control Warnings, trigger "2062_Warning_Data_BTCS_WARNING_WORD_09" bit 8
   2265: 'PS436 RIO2 TANK GROUP PRESURE HIGH HIGH', class Tank Control Warnings, trigger "2062_Warning_Data_BTCS_WARNING_WORD_09" bit 9
   2266: 'PS436 RIO3 TANK GROUP PRESURE HIGH HIGH', class Tank Control Warnings, trigger "2062_Warning_Data_BTCS_WARNING_WORD_09" bit 10
   2267: 'PS436 RIO4 TANK GROUP PRESURE HIGH HIGH', class Tank Control Warnings, trigger "2062_Warning_Data_BTCS_WARNING_WORD_09" bit 11
   2268: 'PS436 RIO5 TANK GROUP PRESURE HIGH HIGH', class Tank Control Warnings, trigger "2062_Warning_Data_BTCS_WARNING_WORD_09" bit 12
   2269: 'PS436 RIO6 TANK GROUP PRESURE HIGH HIGH', class Tank Control Warnings, trigger "2062_Warning_Data_BTCS_WARNING_WORD_09" bit 13
   2270: 'PS436 RIO7 TANK GROUP PRESURE HIGH HIGH', class Tank Control Warnings, trigger "2062_Warning_Data_BTCS_WARNING_WORD_09" bit 14
   2271: 'LS425 1 PORT TANK LEVEL HIGH HIGH', class Tank Control Warnings, trigger "2062_Warning_Data_BTCS_WARNING_WORD_09" bit 15
   2032: 'PT415 RIO1 DECK IG PRESSURE LOW LOW', class Tank Control Alarms, trigger "2060_Alarm_Data_BTCS_ALARM_WORD_03" bit 0
   2033: '', class Tank Control Alarms, trigger "2060_Alarm_Data_BTCS_ALARM_WORD_03" bit 1
   2034: 'PT415 RIO1 DECK IG PRESSURE HGH HIGH', class Tank Control Alarms, trigger "2060_Alarm_Data_BTCS_ALARM_WORD_03" bit 2
   2035: 'PT415 RIO3 DECK IG PRESSURE LOW LOW', class Tank Control Alarms, trigger "2060_Alarm_Data_BTCS_ALARM_WORD_03" bit 3
   2036: 'PT415 RIO3 DECK IG PRESSURE HGH HIGH', class Tank Control Alarms, trigger "2060_Alarm_Data_BTCS_ALARM_WORD_03" bit 4
   2037: 'PT415 RIO4 DECK IG PRESSURE LOW LOW', class Tank Control Alarms, trigger "2060_Alarm_Data_BTCS_ALARM_WORD_03" bit 5
   2038: 'PT415 RIO4 DECK IG PRESSURE HGH HIGH', class Tank Control Alarms, trigger "2060_Alarm_Data_BTCS_ALARM_WORD_03" bit 6
   2039: '', class Tank Control Alarms, trigger "2060_Alarm_Data_BTCS_ALARM_WORD_03" bit 7
   2040: 'CV422 5 STARBOARD GAS to TANK VALVE FAULT', class Tank Control Alarms, trigger "2060_Alarm_Data_BTCS_ALARM_WORD_03" bit 8
   2041: 'CV422 6 PORT GAS to TANK VALVE FAULT', class Tank Control Alarms, trigger "2060_Alarm_Data_BTCS_ALARM_WORD_03" bit 9
   2042: 'CV422 6 STARBOARD GAS to TANK VALVE FAULT', class Tank Control Alarms, trigger "2060_Alarm_Data_BTCS_ALARM_WORD_03" bit 10
   2043: 'CV422 APT GAS to TANK VALVE FAULT', class Tank Control Alarms, trigger "2060_Alarm_Data_BTCS_ALARM_WORD_03" bit 11
   2044: '', class Tank Control Alarms, trigger "2060_Alarm_Data_BTCS_ALARM_WORD_03" bit 12
   2045: '', class Tank Control Alarms, trigger "2060_Alarm_Data_BTCS_ALARM_WORD_03" bit 13
   2046: '', class Tank Control Alarms, trigger "2060_Alarm_Data_BTCS_ALARM_WORD_03" bit 14
   2047: '', class Tank Control Alarms, trigger "2060_Alarm_Data_BTCS_ALARM_WORD_03" bit 15
   2048: '', class Tank Control Alarms, trigger "2060_Alarm_Data_BTCS_ALARM_WORD_04" bit 0
   2049: '', class Tank Control Alarms, trigger "2060_Alarm_Data_BTCS_ALARM_WORD_04" bit 1
   2050: '', class Tank Control Alarms, trigger "2060_Alarm_Data_BTCS_ALARM_WORD_04" bit 2
   2051: '', class Tank Control Alarms, trigger "2060_Alarm_Data_BTCS_ALARM_WORD_04" bit 3
   2052: '', class Tank Control Alarms, trigger "2060_Alarm_Data_BTCS_ALARM_WORD_04" bit 4
   2053: '', class Tank Control Alarms, trigger "2060_Alarm_Data_BTCS_ALARM_WORD_04" bit 5
   2054: '', class Tank Control Alarms, trigger "2060_Alarm_Data_BTCS_ALARM_WORD_04" bit 6
   2055: '', class Tank Control Alarms, trigger "2060_Alarm_Data_BTCS_ALARM_WORD_04" bit 7
   2056: 'PT415 RIO5 DECK IG PRESSURE LOW LOW', class Tank Control Alarms, trigger "2060_Alarm_Data_BTCS_ALARM_WORD_04" bit 8
   2057: 'PT415 RIO5 DECK IG PRESSURE HGH HIGH', class Tank Control Alarms, trigger "2060_Alarm_Data_BTCS_ALARM_WORD_04" bit 9
   2058: 'PT415 RIO6 DECK IG PRESSURE LOW LOW', class Tank Control Alarms, trigger "2060_Alarm_Data_BTCS_ALARM_WORD_04" bit 10
   2059: 'PT415 RIO6 DECK IG PRESSURE HGH HIGH', class Tank Control Alarms, trigger "2060_Alarm_Data_BTCS_ALARM_WORD_04" bit 11
   2060: 'PT415 RIO7 DECK IG PRESSURE LOW LOW', class Tank Control Alarms, trigger "2060_Alarm_Data_BTCS_ALARM_WORD_04" bit 12
   2061: 'PT415 RIO7 DECK IG PRESSURE HIGH HIGH', class Tank Control Alarms, trigger "2060_Alarm_Data_BTCS_ALARM_WORD_04" bit 13
   2062: '', class Tank Control Alarms, trigger "2060_Alarm_Data_BTCS_ALARM_WORD_04" bit 14
   2063: '', class Tank Control Alarms, trigger "2060_Alarm_Data_BTCS_ALARM_WORD_04" bit 15
   2272: 'LT422 4 STARBOARD TANK LEVEL HIGH', class Tank Control Warnings, trigger "2062_Warning_Data_BTCS_WARNING_WORD_10" bit 0
   2273: 'LT422 4 STARBOARD TANK LEVEL LOW', class Tank Control Warnings, trigger "2062_Warning_Data_BTCS_WARNING_WORD_10" bit 1
   2274: 'LT422 5 PORT TANK LEVEL HIGH', class Tank Control Warnings, trigger "2062_Warning_Data_BTCS_WARNING_WORD_10" bit 2
   2275: 'LT422 5 PORT TANK LEVEL LOW', class Tank Control Warnings, trigger "2062_Warning_Data_BTCS_WARNING_WORD_10" bit 3
   2276: 'LT422 5 STARBOARD TANK LEVEL HIGH', class Tank Control Warnings, trigger "2062_Warning_Data_BTCS_WARNING_WORD_10" bit 4
   2277: 'LT422 5 STARBOARD TANK LEVEL LOW', class Tank Control Warnings, trigger "2062_Warning_Data_BTCS_WARNING_WORD_10" bit 5
   2278: 'LT422 6 PORT TANK LEVEL HIGH', class Tank Control Warnings, trigger "2062_Warning_Data_BTCS_WARNING_WORD_10" bit 6
   2279: 'LT422 6 PORT TANK LEVEL LOW', class Tank Control Warnings, trigger "2062_Warning_Data_BTCS_WARNING_WORD_10" bit 7
   2280: 'LT422 2 STARBOARD TANK LEVEL HIGH', class Tank Control Warnings, trigger "2062_Warning_Data_BTCS_WARNING_WORD_10" bit 8
   2281: 'LT422 2 STARBOARD TANK LEVEL LOW', class Tank Control Warnings, trigger "2062_Warning_Data_BTCS_WARNING_WORD_10" bit 9
   2282: 'LT422 3 PORT TANK LEVEL HIGH', class Tank Control Warnings, trigger "2062_Warning_Data_BTCS_WARNING_WORD_10" bit 10
   2283: 'LT422 3 PORT TANK LEVEL LOW', class Tank Control Warnings, trigger "2062_Warning_Data_BTCS_WARNING_WORD_10" bit 11
   2284: 'LT422 3 STARBOARD TANK LEVEL HIGH', class Tank Control Warnings, trigger "2062_Warning_Data_BTCS_WARNING_WORD_10" bit 12
   2285: 'LT422 3 STARBOARD TANK LEVEL LOW', class Tank Control Warnings, trigger "2062_Warning_Data_BTCS_WARNING_WORD_10" bit 13
   2286: 'LT422 4 PORT TANK LEVEL HIGH', class Tank Control Warnings, trigger "2062_Warning_Data_BTCS_WARNING_WORD_10" bit 14
   2287: 'LT422 4 PORT TANK LEVEL LOW', class Tank Control Warnings, trigger "2062_Warning_Data_BTCS_WARNING_WORD_10" bit 15
   2288: 'TT426 2S BWT TEMP OUT OF RANGE', class Tank Control Warnings, trigger "2062_Warning_Data_BTCS_WARNING_WORD_11" bit 0
   2289: 'TT426 3P BWT TEMP OUT OF RANGE', class Tank Control Warnings, trigger "2062_Warning_Data_BTCS_WARNING_WORD_11" bit 1